REGION Network 4: Sumowanie parametrów z każdego z ostatnich 7. dni
   // Sumowane jest maksymalnie 16 parametrów z każdego dnia. Wyjątkiem są parametry dla których jakikolwiek parametr nie został odczytany (nie mieści się w wymaganym zakresie).
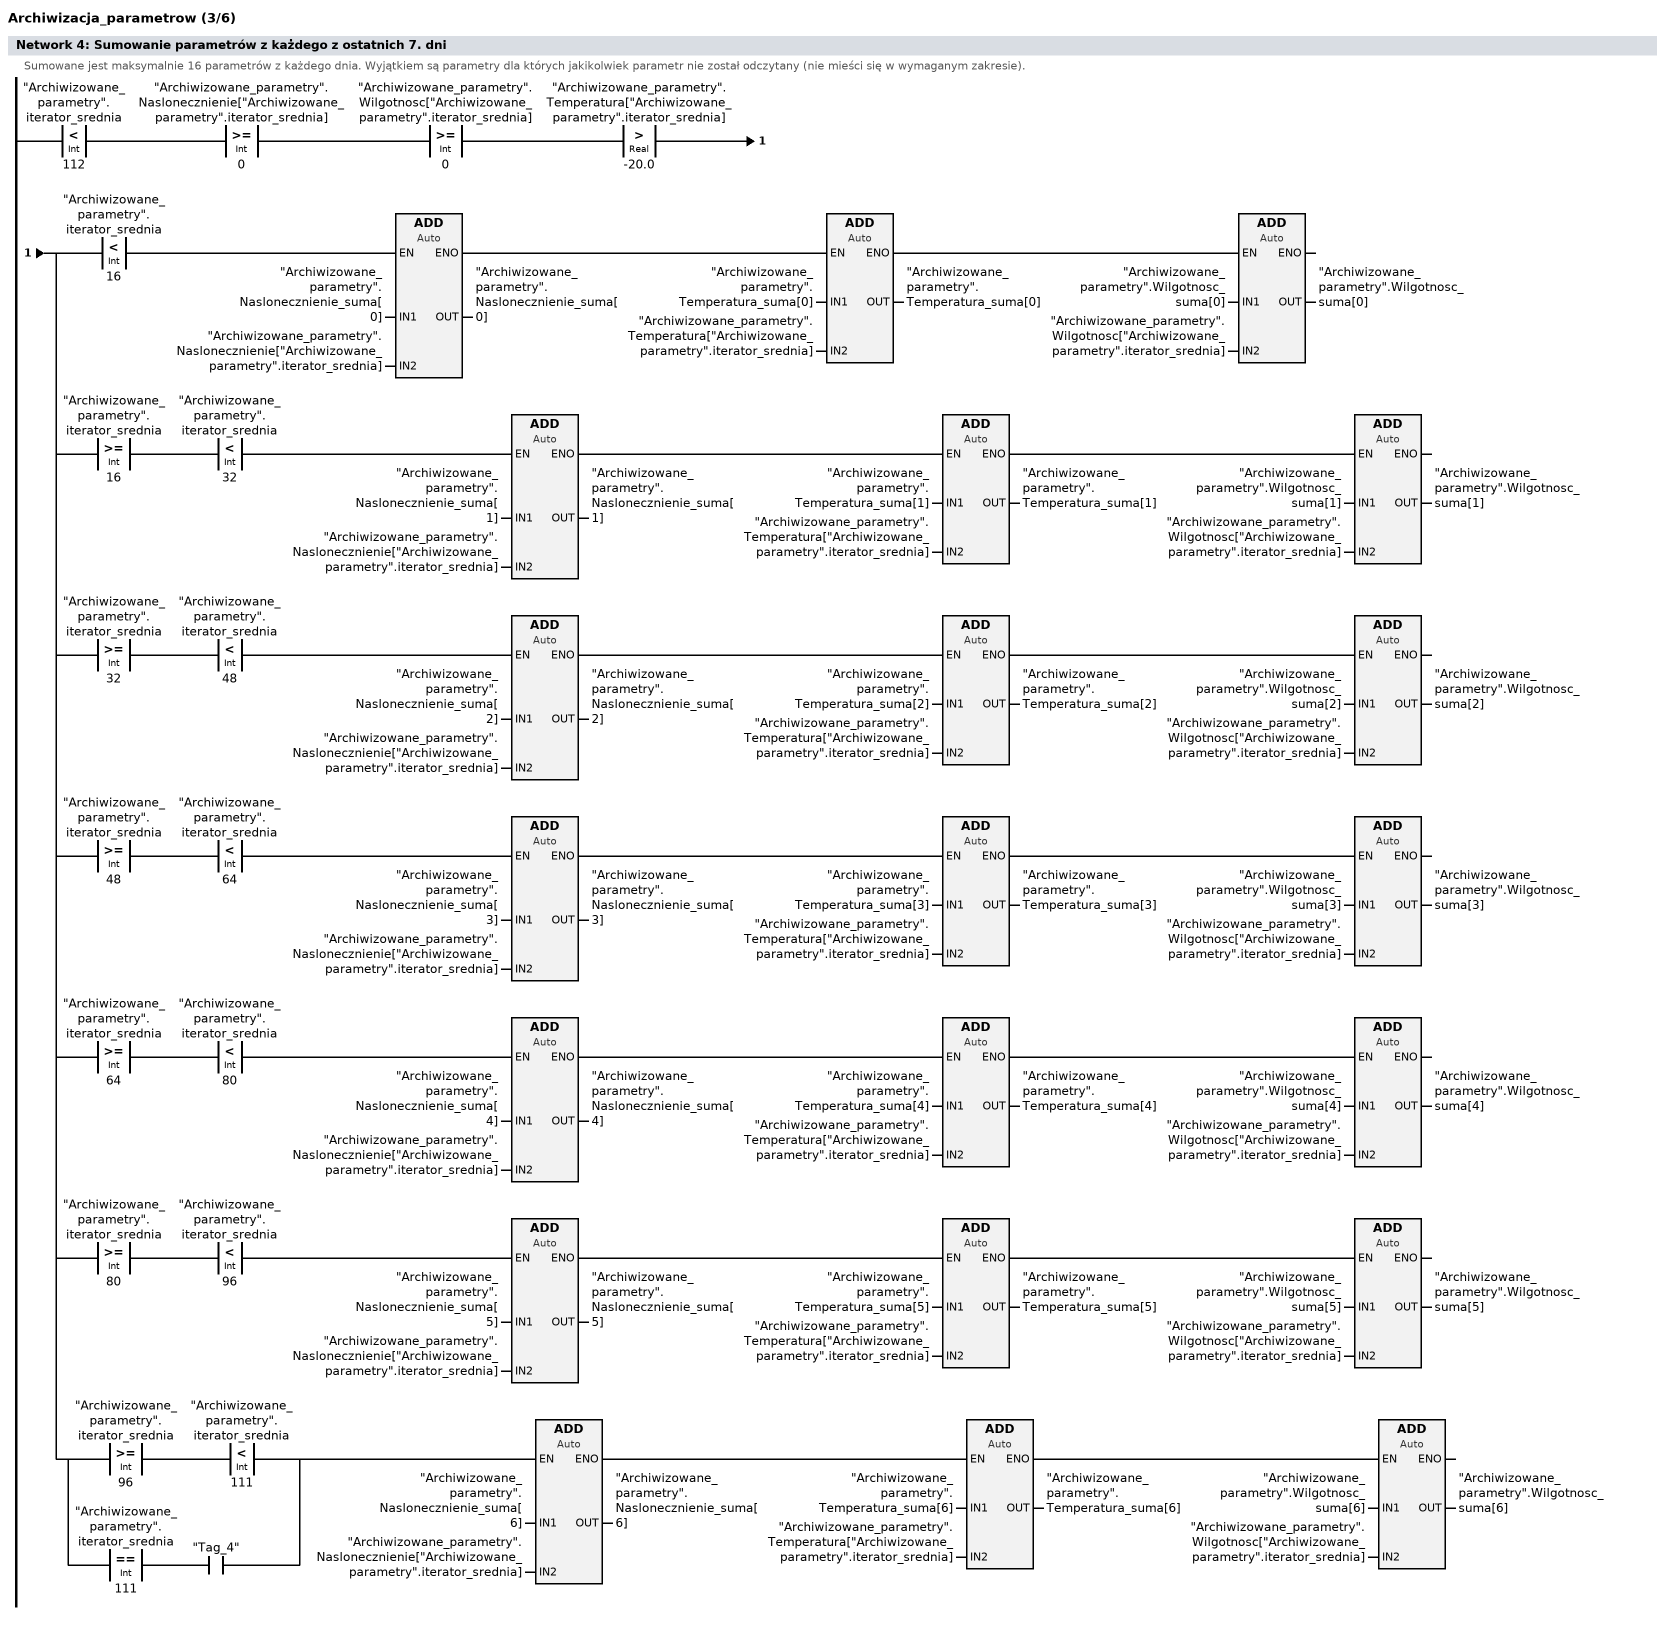
   RUNG wire#powerrail
      { S7_Templates := "SrcType := Int" } LT_Contact(in1 := "Archiwizowane_parametry".iterator_srednia, in2 := 112)
      { S7_Templates := "SrcType := Int" } GE_Contact(in1 := "Archiwizowane_parametry".Naslonecznienie["Archiwizowane_parametry".iterator_srednia], in2 := 0)
      { S7_Templates := "SrcType := Int" } GE_Contact(in1 := "Archiwizowane_parametry".Wilgotnosc["Archiwizowane_parametry".iterator_srednia], in2 := 0)
      { S7_Templates := "SrcType := Real" } GT_Contact(in1 := "Archiwizowane_parametry".Temperatura["Archiwizowane_parametry".iterator_srednia], in2 := -20.0)
      wire#w1
      { S7_Templates := "SrcType := Int" } LT_Contact(in1 := "Archiwizowane_parametry".iterator_srednia, in2 := 16)
      { S7_GenerateENO := "TRUE" } Add(in1 := "Archiwizowane_parametry".Naslonecznienie_suma[0], in2 := "Archiwizowane_parametry".Naslonecznienie["Archiwizowane_parametry".iterator_srednia], out => "Archiwizowane_parametry".Naslonecznienie_suma[0])
      { S7_GenerateENO := "TRUE" } Add(in1 := "Archiwizowane_parametry".Temperatura_suma[0], in2 := "Archiwizowane_parametry".Temperatura["Archiwizowane_parametry".iterator_srednia], out => "Archiwizowane_parametry".Temperatura_suma[0])
      { S7_GenerateENO := "TRUE" } Add(in1 := "Archiwizowane_parametry".Wilgotnosc_suma[0], in2 := "Archiwizowane_parametry".Wilgotnosc["Archiwizowane_parametry".iterator_srednia], out => "Archiwizowane_parametry".Wilgotnosc_suma[0])
   END_RUNG
   RUNG wire#w1
      { S7_Templates := "SrcType := Int" } GE_Contact(in1 := "Archiwizowane_parametry".iterator_srednia, in2 := 16)
      { S7_Templates := "SrcType := Int" } LT_Contact(in1 := "Archiwizowane_parametry".iterator_srednia, in2 := 32)
      { S7_GenerateENO := "TRUE" } Add(in1 := "Archiwizowane_parametry".Naslonecznienie_suma[1], in2 := "Archiwizowane_parametry".Naslonecznienie["Archiwizowane_parametry".iterator_srednia], out => "Archiwizowane_parametry".Naslonecznienie_suma[1])
      { S7_GenerateENO := "TRUE" } Add(in1 := "Archiwizowane_parametry".Temperatura_suma[1], in2 := "Archiwizowane_parametry".Temperatura["Archiwizowane_parametry".iterator_srednia], out => "Archiwizowane_parametry".Temperatura_suma[1])
      { S7_GenerateENO := "TRUE" } Add(in1 := "Archiwizowane_parametry".Wilgotnosc_suma[1], in2 := "Archiwizowane_parametry".Wilgotnosc["Archiwizowane_parametry".iterator_srednia], out => "Archiwizowane_parametry".Wilgotnosc_suma[1])
   END_RUNG
   RUNG wire#w1
      { S7_Templates := "SrcType := Int" } GE_Contact(in1 := "Archiwizowane_parametry".iterator_srednia, in2 := 32)
      { S7_Templates := "SrcType := Int" } LT_Contact(in1 := "Archiwizowane_parametry".iterator_srednia, in2 := 48)
      { S7_GenerateENO := "TRUE" } Add(in1 := "Archiwizowane_parametry".Naslonecznienie_suma[2], in2 := "Archiwizowane_parametry".Naslonecznienie["Archiwizowane_parametry".iterator_srednia], out => "Archiwizowane_parametry".Naslonecznienie_suma[2])
      { S7_GenerateENO := "TRUE" } Add(in1 := "Archiwizowane_parametry".Temperatura_suma[2], in2 := "Archiwizowane_parametry".Temperatura["Archiwizowane_parametry".iterator_srednia], out => "Archiwizowane_parametry".Temperatura_suma[2])
      { S7_GenerateENO := "TRUE" } Add(in1 := "Archiwizowane_parametry".Wilgotnosc_suma[2], in2 := "Archiwizowane_parametry".Wilgotnosc["Archiwizowane_parametry".iterator_srednia], out => "Archiwizowane_parametry".Wilgotnosc_suma[2])
   END_RUNG
   RUNG wire#w1
      { S7_Templates := "SrcType := Int" } GE_Contact(in1 := "Archiwizowane_parametry".iterator_srednia, in2 := 48)
      { S7_Templates := "SrcType := Int" } LT_Contact(in1 := "Archiwizowane_parametry".iterator_srednia, in2 := 64)
      { S7_GenerateENO := "TRUE" } Add(in1 := "Archiwizowane_parametry".Naslonecznienie_suma[3], in2 := "Archiwizowane_parametry".Naslonecznienie["Archiwizowane_parametry".iterator_srednia], out => "Archiwizowane_parametry".Naslonecznienie_suma[3])
      { S7_GenerateENO := "TRUE" } Add(in1 := "Archiwizowane_parametry".Temperatura_suma[3], in2 := "Archiwizowane_parametry".Temperatura["Archiwizowane_parametry".iterator_srednia], out => "Archiwizowane_parametry".Temperatura_suma[3])
      { S7_GenerateENO := "TRUE" } Add(in1 := "Archiwizowane_parametry".Wilgotnosc_suma[3], in2 := "Archiwizowane_parametry".Wilgotnosc["Archiwizowane_parametry".iterator_srednia], out => "Archiwizowane_parametry".Wilgotnosc_suma[3])
   END_RUNG
   RUNG wire#w1
      { S7_Templates := "SrcType := Int" } GE_Contact(in1 := "Archiwizowane_parametry".iterator_srednia, in2 := 64)
      { S7_Templates := "SrcType := Int" } LT_Contact(in1 := "Archiwizowane_parametry".iterator_srednia, in2 := 80)
      { S7_GenerateENO := "TRUE" } Add(in1 := "Archiwizowane_parametry".Naslonecznienie_suma[4], in2 := "Archiwizowane_parametry".Naslonecznienie["Archiwizowane_parametry".iterator_srednia], out => "Archiwizowane_parametry".Naslonecznienie_suma[4])
      { S7_GenerateENO := "TRUE" } Add(in1 := "Archiwizowane_parametry".Temperatura_suma[4], in2 := "Archiwizowane_parametry".Temperatura["Archiwizowane_parametry".iterator_srednia], out => "Archiwizowane_parametry".Temperatura_suma[4])
      { S7_GenerateENO := "TRUE" } Add(in1 := "Archiwizowane_parametry".Wilgotnosc_suma[4], in2 := "Archiwizowane_parametry".Wilgotnosc["Archiwizowane_parametry".iterator_srednia], out => "Archiwizowane_parametry".Wilgotnosc_suma[4])
   END_RUNG
   RUNG wire#w1
      { S7_Templates := "SrcType := Int" } GE_Contact(in1 := "Archiwizowane_parametry".iterator_srednia, in2 := 80)
      { S7_Templates := "SrcType := Int" } LT_Contact(in1 := "Archiwizowane_parametry".iterator_srednia, in2 := 96)
      { S7_GenerateENO := "TRUE" } Add(in1 := "Archiwizowane_parametry".Naslonecznienie_suma[5], in2 := "Archiwizowane_parametry".Naslonecznienie["Archiwizowane_parametry".iterator_srednia], out => "Archiwizowane_parametry".Naslonecznienie_suma[5])
      { S7_GenerateENO := "TRUE" } Add(in1 := "Archiwizowane_parametry".Temperatura_suma[5], in2 := "Archiwizowane_parametry".Temperatura["Archiwizowane_parametry".iterator_srednia], out => "Archiwizowane_parametry".Temperatura_suma[5])
      { S7_GenerateENO := "TRUE" } Add(in1 := "Archiwizowane_parametry".Wilgotnosc_suma[5], in2 := "Archiwizowane_parametry".Wilgotnosc["Archiwizowane_parametry".iterator_srednia], out => "Archiwizowane_parametry".Wilgotnosc_suma[5])
   END_RUNG
   RUNG wire#w1
      { S7_Templates := "SrcType := Int" } GE_Contact(in1 := "Archiwizowane_parametry".iterator_srednia, in2 := 96)
      { S7_Templates := "SrcType := Int" } LT_Contact(in1 := "Archiwizowane_parametry".iterator_srednia, in2 := 111)
      wire#w2
      { S7_GenerateENO := "TRUE" } Add(in1 := "Archiwizowane_parametry".Naslonecznienie_suma[6], in2 := "Archiwizowane_parametry".Naslonecznienie["Archiwizowane_parametry".iterator_srednia], out => "Archiwizowane_parametry".Naslonecznienie_suma[6])
      { S7_GenerateENO := "TRUE" } Add(in1 := "Archiwizowane_parametry".Temperatura_suma[6], in2 := "Archiwizowane_parametry".Temperatura["Archiwizowane_parametry".iterator_srednia], out => "Archiwizowane_parametry".Temperatura_suma[6])
      { S7_GenerateENO := "TRUE" } Add(in1 := "Archiwizowane_parametry".Wilgotnosc_suma[6], in2 := "Archiwizowane_parametry".Wilgotnosc["Archiwizowane_parametry".iterator_srednia], out => "Archiwizowane_parametry".Wilgotnosc_suma[6])
   END_RUNG
   RUNG wire#w1
      { S7_Templates := "SrcType := Int" } EQ_Contact(in1 := "Archiwizowane_parametry".iterator_srednia, in2 := 111)
      Contact( "Tag_4" )
   END_RUNG wire#w2
   // the same network as SCL:
   // ENO of a box is taken as its EN; it also drops when the box reports an error
   #_w1 := ("Archiwizowane_parametry".iterator_srednia < 112) AND ("Archiwizowane_parametry".Naslonecznienie["Archiwizowane_parametry".iterator_srednia] >= 0) AND ("Archiwizowane_parametry".Wilgotnosc["Archiwizowane_parametry".iterator_srednia] >= 0) AND ("Archiwizowane_parametry".Temperatura["Archiwizowane_parametry".iterator_srednia] > (-20.0));
   IF #_w1 AND ("Archiwizowane_parametry".iterator_srednia < 16) THEN
       "Archiwizowane_parametry".Naslonecznienie_suma[0] := "Archiwizowane_parametry".Naslonecznienie_suma[0] + "Archiwizowane_parametry".Naslonecznienie["Archiwizowane_parametry".iterator_srednia];
       "Archiwizowane_parametry".Temperatura_suma[0] := "Archiwizowane_parametry".Temperatura_suma[0] + "Archiwizowane_parametry".Temperatura["Archiwizowane_parametry".iterator_srednia];
       "Archiwizowane_parametry".Wilgotnosc_suma[0] := "Archiwizowane_parametry".Wilgotnosc_suma[0] + "Archiwizowane_parametry".Wilgotnosc["Archiwizowane_parametry".iterator_srednia];
   END_IF;
   IF #_w1 AND ("Archiwizowane_parametry".iterator_srednia >= 16) AND ("Archiwizowane_parametry".iterator_srednia < 32) THEN
       "Archiwizowane_parametry".Naslonecznienie_suma[1] := "Archiwizowane_parametry".Naslonecznienie_suma[1] + "Archiwizowane_parametry".Naslonecznienie["Archiwizowane_parametry".iterator_srednia];
       "Archiwizowane_parametry".Temperatura_suma[1] := "Archiwizowane_parametry".Temperatura_suma[1] + "Archiwizowane_parametry".Temperatura["Archiwizowane_parametry".iterator_srednia];
       "Archiwizowane_parametry".Wilgotnosc_suma[1] := "Archiwizowane_parametry".Wilgotnosc_suma[1] + "Archiwizowane_parametry".Wilgotnosc["Archiwizowane_parametry".iterator_srednia];
   END_IF;
   IF #_w1 AND ("Archiwizowane_parametry".iterator_srednia >= 32) AND ("Archiwizowane_parametry".iterator_srednia < 48) THEN
       "Archiwizowane_parametry".Naslonecznienie_suma[2] := "Archiwizowane_parametry".Naslonecznienie_suma[2] + "Archiwizowane_parametry".Naslonecznienie["Archiwizowane_parametry".iterator_srednia];
       "Archiwizowane_parametry".Temperatura_suma[2] := "Archiwizowane_parametry".Temperatura_suma[2] + "Archiwizowane_parametry".Temperatura["Archiwizowane_parametry".iterator_srednia];
       "Archiwizowane_parametry".Wilgotnosc_suma[2] := "Archiwizowane_parametry".Wilgotnosc_suma[2] + "Archiwizowane_parametry".Wilgotnosc["Archiwizowane_parametry".iterator_srednia];
   END_IF;
   IF #_w1 AND ("Archiwizowane_parametry".iterator_srednia >= 48) AND ("Archiwizowane_parametry".iterator_srednia < 64) THEN
       "Archiwizowane_parametry".Naslonecznienie_suma[3] := "Archiwizowane_parametry".Naslonecznienie_suma[3] + "Archiwizowane_parametry".Naslonecznienie["Archiwizowane_parametry".iterator_srednia];
       "Archiwizowane_parametry".Temperatura_suma[3] := "Archiwizowane_parametry".Temperatura_suma[3] + "Archiwizowane_parametry".Temperatura["Archiwizowane_parametry".iterator_srednia];
       "Archiwizowane_parametry".Wilgotnosc_suma[3] := "Archiwizowane_parametry".Wilgotnosc_suma[3] + "Archiwizowane_parametry".Wilgotnosc["Archiwizowane_parametry".iterator_srednia];
   END_IF;
   IF #_w1 AND ("Archiwizowane_parametry".iterator_srednia >= 64) AND ("Archiwizowane_parametry".iterator_srednia < 80) THEN
       "Archiwizowane_parametry".Naslonecznienie_suma[4] := "Archiwizowane_parametry".Naslonecznienie_suma[4] + "Archiwizowane_parametry".Naslonecznienie["Archiwizowane_parametry".iterator_srednia];
       "Archiwizowane_parametry".Temperatura_suma[4] := "Archiwizowane_parametry".Temperatura_suma[4] + "Archiwizowane_parametry".Temperatura["Archiwizowane_parametry".iterator_srednia];
       "Archiwizowane_parametry".Wilgotnosc_suma[4] := "Archiwizowane_parametry".Wilgotnosc_suma[4] + "Archiwizowane_parametry".Wilgotnosc["Archiwizowane_parametry".iterator_srednia];
   END_IF;
   IF #_w1 AND ("Archiwizowane_parametry".iterator_srednia >= 80) AND ("Archiwizowane_parametry".iterator_srednia < 96) THEN
       "Archiwizowane_parametry".Naslonecznienie_suma[5] := "Archiwizowane_parametry".Naslonecznienie_suma[5] + "Archiwizowane_parametry".Naslonecznienie["Archiwizowane_parametry".iterator_srednia];
       "Archiwizowane_parametry".Temperatura_suma[5] := "Archiwizowane_parametry".Temperatura_suma[5] + "Archiwizowane_parametry".Temperatura["Archiwizowane_parametry".iterator_srednia];
       "Archiwizowane_parametry".Wilgotnosc_suma[5] := "Archiwizowane_parametry".Wilgotnosc_suma[5] + "Archiwizowane_parametry".Wilgotnosc["Archiwizowane_parametry".iterator_srednia];
   END_IF;
   IF #_w1 AND ((("Archiwizowane_parametry".iterator_srednia >= 96) AND ("Archiwizowane_parametry".iterator_srednia < 111)) OR (("Archiwizowane_parametry".iterator_srednia = 111) AND "Tag_4")) THEN
       "Archiwizowane_parametry".Naslonecznienie_suma[6] := "Archiwizowane_parametry".Naslonecznienie_suma[6] + "Archiwizowane_parametry".Naslonecznienie["Archiwizowane_parametry".iterator_srednia];
       "Archiwizowane_parametry".Temperatura_suma[6] := "Archiwizowane_parametry".Temperatura_suma[6] + "Archiwizowane_parametry".Temperatura["Archiwizowane_parametry".iterator_srednia];
       "Archiwizowane_parametry".Wilgotnosc_suma[6] := "Archiwizowane_parametry".Wilgotnosc_suma[6] + "Archiwizowane_parametry".Wilgotnosc["Archiwizowane_parametry".iterator_srednia];
   END_IF;
END_REGION

REGION Network 5: Obliczenie wartości dzielnika
   // Utworzony jest specjalny dzielnik, który co rośnie do takiej wartości, jaka jest liczba parametrów zsumowanych danego dnia.
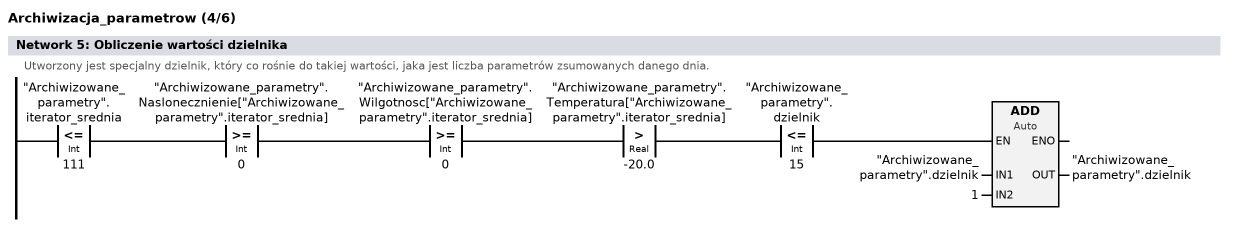
   RUNG wire#powerrail
      { S7_Templates := "SrcType := Int" } LE_Contact(in1 := "Archiwizowane_parametry".iterator_srednia, in2 := 111)
      { S7_Templates := "SrcType := Int" } GE_Contact(in1 := "Archiwizowane_parametry".Naslonecznienie["Archiwizowane_parametry".iterator_srednia], in2 := 0)
      { S7_Templates := "SrcType := Int" } GE_Contact(in1 := "Archiwizowane_parametry".Wilgotnosc["Archiwizowane_parametry".iterator_srednia], in2 := 0)
      { S7_Templates := "SrcType := Real" } GT_Contact(in1 := "Archiwizowane_parametry".Temperatura["Archiwizowane_parametry".iterator_srednia], in2 := -20.0)
      { S7_Templates := "SrcType := Int" } LE_Contact(in1 := "Archiwizowane_parametry".dzielnik, in2 := 15)
      { S7_GenerateENO := "TRUE" } Add(in1 := "Archiwizowane_parametry".dzielnik, in2 := 1, out => "Archiwizowane_parametry".dzielnik)
   END_RUNG
   // the same network as SCL:
   IF ("Archiwizowane_parametry".iterator_srednia <= 111) AND ("Archiwizowane_parametry".Naslonecznienie["Archiwizowane_parametry".iterator_srednia] >= 0) AND ("Archiwizowane_parametry".Wilgotnosc["Archiwizowane_parametry".iterator_srednia] >= 0) AND ("Archiwizowane_parametry".Temperatura["Archiwizowane_parametry".iterator_srednia] > (-20.0)) AND ("Archiwizowane_parametry".dzielnik <= 15) THEN
       "Archiwizowane_parametry".dzielnik := "Archiwizowane_parametry".dzielnik + 1;
   END_IF;
END_REGION

REGION Network 6: Obliczanie średniej parametrów z każdego z ostatnich 7. dni
   // Obliczone wcześniej sumy dzielone są wartość dzielnika, dzięki czemu otrzymywana jest średnia parametrów z każdego z ostatnich 7. dni. Po tym dzielnik jest zerowany.
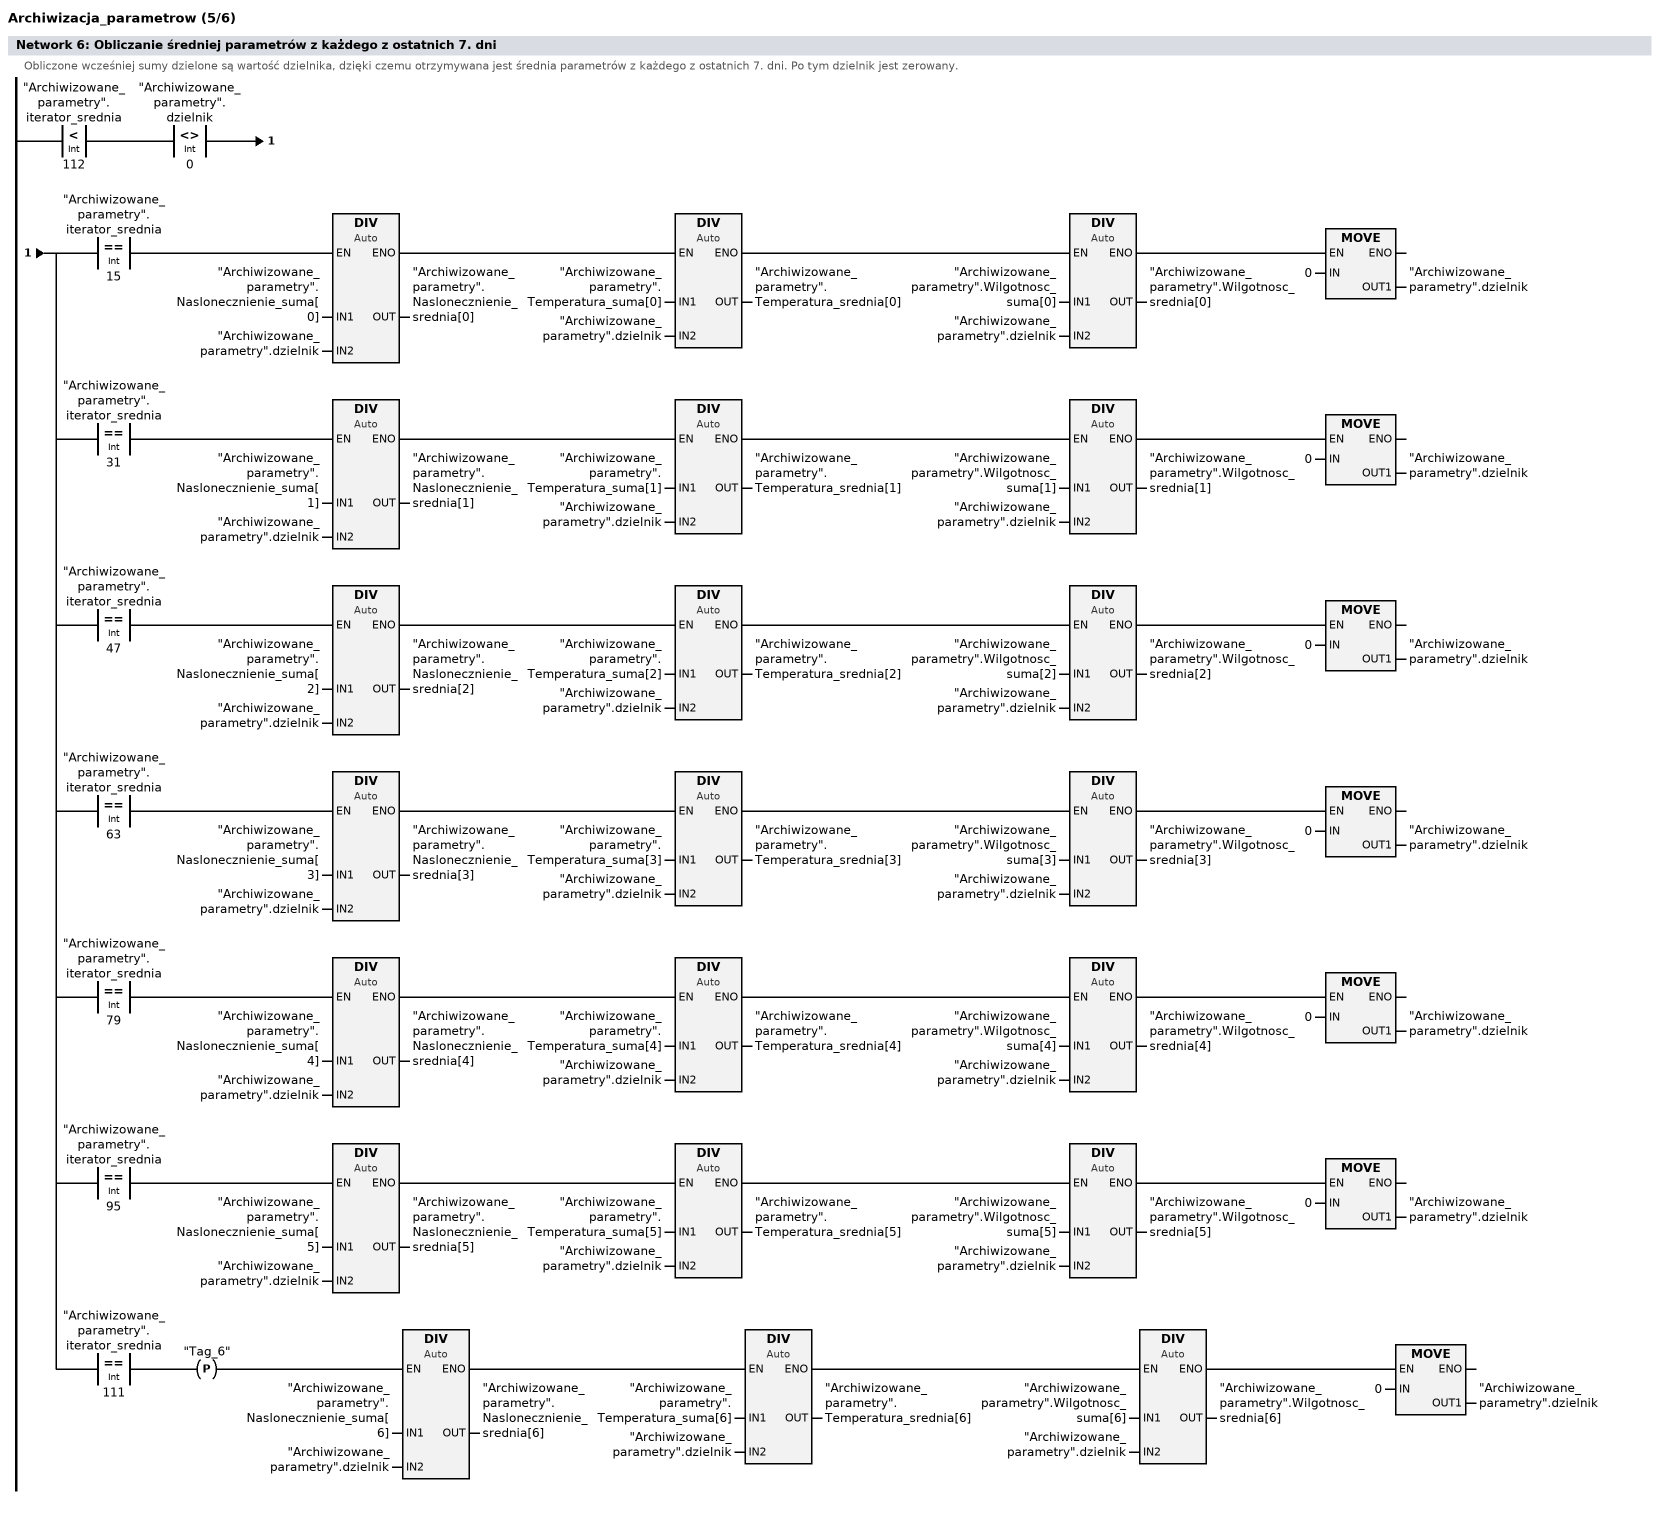
   RUNG wire#powerrail
      { S7_Templates := "SrcType := Int" } LT_Contact(in1 := "Archiwizowane_parametry".iterator_srednia, in2 := 112)
      { S7_Templates := "SrcType := Int" } NE_Contact(in1 := "Archiwizowane_parametry".dzielnik, in2 := 0)
      wire#w1
      { S7_Templates := "SrcType := Int" } EQ_Contact(in1 := "Archiwizowane_parametry".iterator_srednia, in2 := 15)
      Div(in1 := "Archiwizowane_parametry".Naslonecznienie_suma[0], in2 := "Archiwizowane_parametry".dzielnik, out => "Archiwizowane_parametry".Naslonecznienie_srednia[0])
      Div(in1 := "Archiwizowane_parametry".Temperatura_suma[0], in2 := "Archiwizowane_parametry".dzielnik, out => "Archiwizowane_parametry".Temperatura_srednia[0])
      Div(in1 := "Archiwizowane_parametry".Wilgotnosc_suma[0], in2 := "Archiwizowane_parametry".dzielnik, out => "Archiwizowane_parametry".Wilgotnosc_srednia[0])
      Move(in := 0, out1 => "Archiwizowane_parametry".dzielnik)
   END_RUNG
   RUNG wire#w1
      { S7_Templates := "SrcType := Int" } EQ_Contact(in1 := "Archiwizowane_parametry".iterator_srednia, in2 := 31)
      Div(in1 := "Archiwizowane_parametry".Naslonecznienie_suma[1], in2 := "Archiwizowane_parametry".dzielnik, out => "Archiwizowane_parametry".Naslonecznienie_srednia[1])
      Div(in1 := "Archiwizowane_parametry".Temperatura_suma[1], in2 := "Archiwizowane_parametry".dzielnik, out => "Archiwizowane_parametry".Temperatura_srednia[1])
      Div(in1 := "Archiwizowane_parametry".Wilgotnosc_suma[1], in2 := "Archiwizowane_parametry".dzielnik, out => "Archiwizowane_parametry".Wilgotnosc_srednia[1])
      Move(in := 0, out1 => "Archiwizowane_parametry".dzielnik)
   END_RUNG
   RUNG wire#w1
      { S7_Templates := "SrcType := Int" } EQ_Contact(in1 := "Archiwizowane_parametry".iterator_srednia, in2 := 47)
      Div(in1 := "Archiwizowane_parametry".Naslonecznienie_suma[2], in2 := "Archiwizowane_parametry".dzielnik, out => "Archiwizowane_parametry".Naslonecznienie_srednia[2])
      Div(in1 := "Archiwizowane_parametry".Temperatura_suma[2], in2 := "Archiwizowane_parametry".dzielnik, out => "Archiwizowane_parametry".Temperatura_srednia[2])
      Div(in1 := "Archiwizowane_parametry".Wilgotnosc_suma[2], in2 := "Archiwizowane_parametry".dzielnik, out => "Archiwizowane_parametry".Wilgotnosc_srednia[2])
      Move(in := 0, out1 => "Archiwizowane_parametry".dzielnik)
   END_RUNG
   RUNG wire#w1
      { S7_Templates := "SrcType := Int" } EQ_Contact(in1 := "Archiwizowane_parametry".iterator_srednia, in2 := 63)
      Div(in1 := "Archiwizowane_parametry".Naslonecznienie_suma[3], in2 := "Archiwizowane_parametry".dzielnik, out => "Archiwizowane_parametry".Naslonecznienie_srednia[3])
      Div(in1 := "Archiwizowane_parametry".Temperatura_suma[3], in2 := "Archiwizowane_parametry".dzielnik, out => "Archiwizowane_parametry".Temperatura_srednia[3])
      Div(in1 := "Archiwizowane_parametry".Wilgotnosc_suma[3], in2 := "Archiwizowane_parametry".dzielnik, out => "Archiwizowane_parametry".Wilgotnosc_srednia[3])
      Move(in := 0, out1 => "Archiwizowane_parametry".dzielnik)
   END_RUNG
   RUNG wire#w1
      { S7_Templates := "SrcType := Int" } EQ_Contact(in1 := "Archiwizowane_parametry".iterator_srednia, in2 := 79)
      Div(in1 := "Archiwizowane_parametry".Naslonecznienie_suma[4], in2 := "Archiwizowane_parametry".dzielnik, out => "Archiwizowane_parametry".Naslonecznienie_srednia[4])
      Div(in1 := "Archiwizowane_parametry".Temperatura_suma[4], in2 := "Archiwizowane_parametry".dzielnik, out => "Archiwizowane_parametry".Temperatura_srednia[4])
      Div(in1 := "Archiwizowane_parametry".Wilgotnosc_suma[4], in2 := "Archiwizowane_parametry".dzielnik, out => "Archiwizowane_parametry".Wilgotnosc_srednia[4])
      Move(in := 0, out1 => "Archiwizowane_parametry".dzielnik)
   END_RUNG
   RUNG wire#w1
      { S7_Templates := "SrcType := Int" } EQ_Contact(in1 := "Archiwizowane_parametry".iterator_srednia, in2 := 95)
      Div(in1 := "Archiwizowane_parametry".Naslonecznienie_suma[5], in2 := "Archiwizowane_parametry".dzielnik, out => "Archiwizowane_parametry".Naslonecznienie_srednia[5])
      Div(in1 := "Archiwizowane_parametry".Temperatura_suma[5], in2 := "Archiwizowane_parametry".dzielnik, out => "Archiwizowane_parametry".Temperatura_srednia[5])
      Div(in1 := "Archiwizowane_parametry".Wilgotnosc_suma[5], in2 := "Archiwizowane_parametry".dzielnik, out => "Archiwizowane_parametry".Wilgotnosc_srednia[5])
      Move(in := 0, out1 => "Archiwizowane_parametry".dzielnik)
   END_RUNG
   RUNG wire#w1
      { S7_Templates := "SrcType := Int" } EQ_Contact(in1 := "Archiwizowane_parametry".iterator_srednia, in2 := 111)
      P_Trig( "Tag_6" )
      Div(in1 := "Archiwizowane_parametry".Naslonecznienie_suma[6], in2 := "Archiwizowane_parametry".dzielnik, out => "Archiwizowane_parametry".Naslonecznienie_srednia[6])
      Div(in1 := "Archiwizowane_parametry".Temperatura_suma[6], in2 := "Archiwizowane_parametry".dzielnik, out => "Archiwizowane_parametry".Temperatura_srednia[6])
      Div(in1 := "Archiwizowane_parametry".Wilgotnosc_suma[6], in2 := "Archiwizowane_parametry".dzielnik, out => "Archiwizowane_parametry".Wilgotnosc_srednia[6])
      Move(in := 0, out1 => "Archiwizowane_parametry".dzielnik)
   END_RUNG
   // the same network as SCL:
   #_w1 := ("Archiwizowane_parametry".iterator_srednia < 112) AND ("Archiwizowane_parametry".dzielnik <> 0);
   IF #_w1 AND ("Archiwizowane_parametry".iterator_srednia = 15) THEN
       "Archiwizowane_parametry".Naslonecznienie_srednia[0] := "Archiwizowane_parametry".Naslonecznienie_suma[0] / "Archiwizowane_parametry".dzielnik;
       "Archiwizowane_parametry".Temperatura_srednia[0] := "Archiwizowane_parametry".Temperatura_suma[0] / "Archiwizowane_parametry".dzielnik;
       "Archiwizowane_parametry".Wilgotnosc_srednia[0] := "Archiwizowane_parametry".Wilgotnosc_suma[0] / "Archiwizowane_parametry".dzielnik;
       "Archiwizowane_parametry".dzielnik := 0;
   END_IF;
   IF #_w1 AND ("Archiwizowane_parametry".iterator_srednia = 31) THEN
       "Archiwizowane_parametry".Naslonecznienie_srednia[1] := "Archiwizowane_parametry".Naslonecznienie_suma[1] / "Archiwizowane_parametry".dzielnik;
       "Archiwizowane_parametry".Temperatura_srednia[1] := "Archiwizowane_parametry".Temperatura_suma[1] / "Archiwizowane_parametry".dzielnik;
       "Archiwizowane_parametry".Wilgotnosc_srednia[1] := "Archiwizowane_parametry".Wilgotnosc_suma[1] / "Archiwizowane_parametry".dzielnik;
       "Archiwizowane_parametry".dzielnik := 0;
   END_IF;
   IF #_w1 AND ("Archiwizowane_parametry".iterator_srednia = 47) THEN
       "Archiwizowane_parametry".Naslonecznienie_srednia[2] := "Archiwizowane_parametry".Naslonecznienie_suma[2] / "Archiwizowane_parametry".dzielnik;
       "Archiwizowane_parametry".Temperatura_srednia[2] := "Archiwizowane_parametry".Temperatura_suma[2] / "Archiwizowane_parametry".dzielnik;
       "Archiwizowane_parametry".Wilgotnosc_srednia[2] := "Archiwizowane_parametry".Wilgotnosc_suma[2] / "Archiwizowane_parametry".dzielnik;
       "Archiwizowane_parametry".dzielnik := 0;
   END_IF;
   IF #_w1 AND ("Archiwizowane_parametry".iterator_srednia = 63) THEN
       "Archiwizowane_parametry".Naslonecznienie_srednia[3] := "Archiwizowane_parametry".Naslonecznienie_suma[3] / "Archiwizowane_parametry".dzielnik;
       "Archiwizowane_parametry".Temperatura_srednia[3] := "Archiwizowane_parametry".Temperatura_suma[3] / "Archiwizowane_parametry".dzielnik;
       "Archiwizowane_parametry".Wilgotnosc_srednia[3] := "Archiwizowane_parametry".Wilgotnosc_suma[3] / "Archiwizowane_parametry".dzielnik;
       "Archiwizowane_parametry".dzielnik := 0;
   END_IF;
   IF #_w1 AND ("Archiwizowane_parametry".iterator_srednia = 79) THEN
       "Archiwizowane_parametry".Naslonecznienie_srednia[4] := "Archiwizowane_parametry".Naslonecznienie_suma[4] / "Archiwizowane_parametry".dzielnik;
       "Archiwizowane_parametry".Temperatura_srednia[4] := "Archiwizowane_parametry".Temperatura_suma[4] / "Archiwizowane_parametry".dzielnik;
       "Archiwizowane_parametry".Wilgotnosc_srednia[4] := "Archiwizowane_parametry".Wilgotnosc_suma[4] / "Archiwizowane_parametry".dzielnik;
       "Archiwizowane_parametry".dzielnik := 0;
   END_IF;
   IF #_w1 AND ("Archiwizowane_parametry".iterator_srednia = 95) THEN
       "Archiwizowane_parametry".Naslonecznienie_srednia[5] := "Archiwizowane_parametry".Naslonecznienie_suma[5] / "Archiwizowane_parametry".dzielnik;
       "Archiwizowane_parametry".Temperatura_srednia[5] := "Archiwizowane_parametry".Temperatura_suma[5] / "Archiwizowane_parametry".dzielnik;
       "Archiwizowane_parametry".Wilgotnosc_srednia[5] := "Archiwizowane_parametry".Wilgotnosc_suma[5] / "Archiwizowane_parametry".dzielnik;
       "Archiwizowane_parametry".dzielnik := 0;
   END_IF;
   #_w2 := #_w1 AND ("Archiwizowane_parametry".iterator_srednia = 111);
   #_w3 := #_w2 AND NOT "Tag_6";   // rising edge
   "Tag_6" := #_w2;
   IF #_w3 THEN
       "Archiwizowane_parametry".Naslonecznienie_srednia[6] := "Archiwizowane_parametry".Naslonecznienie_suma[6] / "Archiwizowane_parametry".dzielnik;
       "Archiwizowane_parametry".Temperatura_srednia[6] := "Archiwizowane_parametry".Temperatura_suma[6] / "Archiwizowane_parametry".dzielnik;
       "Archiwizowane_parametry".Wilgotnosc_srednia[6] := "Archiwizowane_parametry".Wilgotnosc_suma[6] / "Archiwizowane_parametry".dzielnik;
       "Archiwizowane_parametry".dzielnik := 0;
   END_IF;
END_REGION

REGION Network 7: Zwiększanie wartości iteratora używanego do obliczania średniej